// Mitsubishi GX Works2 project: 30国轩预化成10.29,排队位置优化   PLC: Q10UDEH

TYPE ConveyorIO : STRUCT
  xUnloadCCW : BOOL;  (* 下料为反转 *)
  xUnloadAlarm : BOOL;  (* 下料报警 *)
  xUnload : BOOL;  (* 下料请求 *)
  xPutInto : BOOL;  (* 线体直接投入物料 *)
  xNotArriveAlarm : BOOL;  (* 未到达报警 *)
  xNextRun : BOOL;  (* 下段线体运行 *)
  xMotorCW : BOOL;  (* 电机正转 *)
  xMotorCCW : BOOL;  (* 电机反转 *)
  xManual : BOOL;  (* 手动 *)
  xloadCCW : BOOL;  (* 上料为反转 *)
  xLimitAlarrm : BOOL;  (* 限位报警 *)
  xLoad : BOOL;  (* 上料请求 *)
  xForward : BOOL;  (* 正转手动 *)
  xEmpty : BOOL;  (* 线体状态为空 *)
  xCWPresent : BOOL;  (* 正转检测有无传感器 *)
  xCCWPresent : BOOL;  (* 反转检测有无传感器 *)
  xBusy : BOOL;  (* 工作中 *)
  xBackward : BOOL;  (* 反转手动 *)
  xAuto : BOOL;  (* 自动 *)
  xPosLimit : BOOL;  (* 正限位 *)
  xNegLimit : BOOL;  (* 负限位 *)
  xOverWidthAlarm : BOOL;  (* 超宽报警 *)
  xError : BOOL;  (* 报警 *)
  iProductCategoryIn : INT;  (* 产品类型输入 *)
  iProductCategory : INT;  (* 产品类型记录 *)
  iProductCategoryOut : INT;  (* 产品类型输出 *)
  diDeviceID : DINT;  (* 设备编号 *)
  tUnloadAlarmDelay : TIME;  (* 下料报警时间设置 *)
  tLoadDelay : TIME;  (* 上料延时设置 *)
  xSizeDeficientDetect : BOOL;  (* 尺寸缺陷检测 *)
  xZoneClear : BOOL;  (* 初始化线体清除 *)
  tZoneClearTime : TIME;  (* 初始化线体清除时间 *)
  iTaskIDIn : INT;  (* 产品类型输入 *)
  iTaskID : INT;  (* 产品类型记录 *)
  iTaskIDOut : INT;  (* 产品类型输出 *)
  diDesConveyorIn : DINT;  (* 产品类型输入 *)
  diDesConveyor : DINT;  (* 产品类型记录 *)
  diDesConveyorOut : DINT;  (* 产品类型输出 *)
END_STRUCT END_TYPE

TYPE ShuttleCarIO : STRUCT
  xReady : BOOL;  (* 准备就绪 *)
  xForward : BOOL;  (* 正转 *)
  xBackward : BOOL;  (* 反转 *)
  iCurrentPos : INT;  (* 当前位置 *)
  iDestinationPos : INT;  (* 目标位置 *)
  xCW : BOOL;  (* 正转输出 *)
  xCCW : BOOL;  (* 反转输出 *)
  xBrake : BOOL;  (* 刹车 *)
  xHomeSwitch : BOOL;  (* 零位接近开关 *)
  xPosLimit : BOOL;  (* 正限位 *)
  xNegLimit : BOOL;  (* 负限位 *)
  xMDIExe : BOOL;  (* MDI开始 *)
  xMDIDone : BOOL;  (* MDI 完成 *)
  xPassLimit : BOOL;  (* 限位屏蔽 *)
  xPosLimitCatch : BOOL;  (* 正限位捕捉 *)
  xNegLimitCatch : BOOL;  (* 负限位捕捉 *)
  xHomeExe : BOOL;  (* 开始寻零 *)
  xHomeDone : BOOL;  (* 寻零完成 *)
  xHomeBusy : BOOL;  (* 寻零中 *)
  xHomeFailed : BOOL;  (* 寻零失败 *)
  xBusy : BOOL;  (* 工作中 *)
  tArriveDelay : TIME;  (* 到位延时 *)
  xCylinder : BOOL;  (* 气缸控制 *)
  tBrakeDelay : TIME;  (* 抱闸延时 *)
  xPauseRamp : BOOL;  (* 暂停减速斜坡标志位 *)
  xPresentDetect1 : BOOL;  (* 物料有无检测1 *)
  xPresentDetect2 : BOOL;  (* 物料有无检测2 *)
  xOvertimeAlarm : BOOL;  (* 超时报警 *)
  tSetOverTime : TIME;  (* 设置超时时间 *)
  xLooseDetect : BOOL;  (* 松绳检测 *)
  xLooseAlarm : BOOL;  (* 松绳报警 *)
  xArrive : BOOL;  (* 到位信号 *)
  diDeviceID : DINT;  (* 设备编号 *)
  xMoveStep : BOOL;  (* 寸动 *)
  xAdrSwitch : ARRAY [1..8] OF BOOL;  (* 位置开关 *)
END_STRUCT END_TYPE

TYPE SwitchIO : STRUCT
  xLiftCylinderRetractDetect : BOOL;
  xLiftCylinderExtendDetect : BOOL;
  xLiftCylinderRetract : BOOL;
  xLiftCylinderExtend : BOOL;
  xEntryBarCylinderRetract : BOOL;
  xLiftCylinderExtendInit : BOOL;
  xEntryEnable : BOOL;
  xExitEnable : BOOL;
  xExitBarCylinderRetract : BOOL;
  xSwithEnable : BOOL;
  xLiftCylinderRetractButton : BOOL;
  xLiftCylinderExtendButton : BOOL;
  xEntryBarCylinderRetractButton : BOOL;
  xExitBarCylinderRetractButton : BOOL;
  xPutInto : BOOL;  (* 单体复位 *)
  tSetOvertime : TIME;  (* 设定超时报警时间 *)
  xOvertimeAlarm : BOOL;  (* 超时报警 *)
END_STRUCT END_TYPE

TYPE QueueElement : STRUCT
  xCondition : BOOL;
  iPriority : INT;
END_STRUCT END_TYPE

TYPE UConveyorIO : STRUCT
  xLiftCylinderRetractDetect1 : BOOL;
  xLiftCylinderRetractDetect2 : BOOL;
  xLiftCylinderExtendDetect1 : BOOL;
  xLiftCylinderExtendDetect2 : BOOL;
  xLiftCylinderRetract1 : BOOL;
  xLiftCylinderRetract2 : BOOL;
  xLiftCylinderExtend1 : BOOL;
  xLiftCylinderExtend2 : BOOL;
  xExitBarCylinderRetract1 : BOOL;
  xExitBarCylinderRetract2 : BOOL;
  xLiftCylinderExtendInit1 : BOOL;
  xLiftCylinderExtendInit2 : BOOL;
  xEntryEnable1 : BOOL;
  xEntryEnable2 : BOOL;
  xEntryEnable3 : BOOL;
  xExitEnable1 : BOOL;
  xExitEnable2 : BOOL;
  xExitEnable3 : BOOL;
  xPassEnable : BOOL;  (* 直接放行去下段 *)
  xLiftCylinderRetractButton1 : BOOL;
  xLiftCylinderRetractButton2 : BOOL;
  xLiftCylinderExtendButton1 : BOOL;
  xLiftCylinderExtendButton2 : BOOL;
  xExitBarCylinderRetractButton1 : BOOL;
  xExitBarCylinderRetractButton2 : BOOL;
  xPutInto : BOOL;  (* 单体复位 *)
  tSetOvertime : TIME;  (* 设定超时报警时间 *)
  xOvertimeAlarm : BOOL;  (* 超时报警 *)
  iTask : INT;  (* 3个任务 *)
  xBatteryDetect1 : BOOL;  (* 电池检测1 *)
  xBatteryDetect2 : BOOL;  (* 电池检测2 *)
  xBatteryError : BOOL;  (* 空框里有电池错误 *)
END_STRUCT END_TYPE

TYPE FolderIO : STRUCT
  o_xCylinderGrabExtend : BOOL;  (* 气缸夹紧 *)
  o_xCylinderGrabRetract : BOOL;  (* 气缸松开 *)
  i_xCylinderGrabExtendDetect : BOOL;  (* 夹紧检测 *)
  i_xCylinderGrabRetractDetect : BOOL;  (* 松开检测 *)
  o_xCylinderUpExtend : BOOL;  (* 上层伸出 *)
  o_xCylinderUpRetract : BOOL;  (* 上层缩回 *)
  i_xCylinderUpExtendDetect : BOOL;  (* 上层伸出检测 *)
  i_xCylinderUpRetractDetect : BOOL;  (* 上层缩回检测 *)
  o_xCylinderDownExtend : BOOL;  (* 下层伸出 *)
  o_xCylinderDownRetract : BOOL;  (* 下层缩回 *)
  i_xCylinderDownExtendDetect : BOOL;  (* 下层伸出检测 *)
  i_xCylinderDownRetractDetect : BOOL;  (* 下层缩回检测 *)
  i_xExitEnable : BOOL;  (* 下料信号 *)
  i_xEntryEnable : BOOL;  (* 上料信号 *)
  o_xEntryPermit : BOOL;  (* 允许上料 *)
  i_iFloor : INT;  (* 层数 *)
  i_xCylinderGrabExtendButton : BOOL;  (* 气缸夹紧按钮 *)
  i_xCylinderGrabRetractButton : BOOL;  (* 气缸松开按钮 *)
  i_xCylinderUpExtendButton : BOOL;  (* 上层伸出按钮 *)
  i_xCylinderUpRetractButton : BOOL;  (* 上层缩回按钮 *)
  i_xCylinderDownExtendButton : BOOL;  (* 下层伸出按钮 *)
  i_xCylinderDownRetractButton : BOOL;  (* 下层缩回按钮 *)
  o_xDownCylinderError : BOOL;  (* 下层气缸层伸出未到达 *)
  o_xUpCylinderError : BOOL;  (* 上层气缸伸出未到达 *)
  o_xGrabCylinderError : BOOL;  (* 夹紧气缸伸出未到达 *)
  i_tSetOvertime : TIME;  (* 未到达计时 *)
END_STRUCT END_TYPE

TYPE CommunicationIO : STRUCT
  i_iResponsPCPLC : INT;  (* 上位机写入-请求确认 *)
  i_iReadWriteFlagPCPLC : INT;  (* 上位机写入-读写标志位 *)
  i_iTaskProcessFlagPCPLC : INT;  (* 上位机写入-任务处理标志位 *)
  i_iCommandPCPLC : INT;  (* 上位机写入-命令字 *)
  i_iTaskIDPCPLC : INT;  (* 上位机写入-任务号 *)
  i_diDestinationDevicePCPLC : DINT;  (* 上位机写入-目标设备号 *)
  i_iProductIDPCPLC : INT;  (* 上位机写入-框码后4位 *)
  o_iRequestPLCPC : INT;  (* 上位机读取-请求状态 *)
  o_iReadWriteFlagPLCPC : INT;  (* 上位机读取-读写标志位 *)
  o_iDeviceStatusPLCPC : INT;  (* 上位机读取-设备状态 *)
  o_iTaskIDPLCPC : INT;  (* 上位机读取-任务号 *)
  o_iProductIDPLCPC : INT;  (* 上位机读取-框码后4位 *)
  i_iTypeInfoPCPLC : INT;  (* 上位机写入-批次标识，是否同批次 *)
  o_iForceInportPLCPC : INT;  (* 上位机读取-强制入库 *)
  o_iEmptyPLCPC : INT;  (* 上位机读取-有料状态 *)
  o_iFolderNumberPLCPC : INT;  (* 上位机读取-叠盘数量 *)
  i_xExtraCondition : BOOL;  (* 发送请求时的额外条件,比如需要升降到位 *)
  i_xExportConveyor : BOOL;  (* 线体是出库线体还是入库线体 *)
END_STRUCT END_TYPE

TYPE FanucRobotIO : STRUCT
  i_xCMDENBL : BOOL;
  i_xSYSRDY : BOOL;
  i_xPROG_RUN : BOOL;  (* 程序运行中 *)
  i_xPAUSED : BOOL;
  i_xHELD : BOOL;
  i_xFAULT : BOOL;
  i_xATPERCH : BOOL;
  i_xTPENBL : BOOL;
  i_xBATALM : BOOL;
  i_xBUSY : BOOL;  (* 工作中信号 *)
  i_arrxSNO : ARRAY [0..7] OF BOOL;  (* 传回的数据 *)
  i_xSNACK : BOOL;  (* 数据传回校验标志位 *)
  o_xIMSTP : BOOL;
  o_xHOLD : BOOL;
  o_xSFSPD : BOOL;
  o_xCSTOPI : BOOL;
  o_xRESET : BOOL;
  o_xSTART : BOOL;
  o_xENBL : BOOL;
  o_iPNS : INT;  (* 发给他的动作编号 *)
  o_xPNSTROBE : BOOL;  (* 传递动作编号标志位 *)
  o_xPROD_START : BOOL;  (* 启动信号，下降沿开动 *)
  o_xREMOTE : BOOL;  (* 远程模式开启 *)
  i_xCommandStart : BOOL;  (* 启动 *)
  i_iMotionNumber : INT;  (* 我程序给的动作编号 *)
  o_xPNSFailed : BOOL;  (* 程序号传输错误 *)
  o_uiOffset_X : INT;  (* X轴偏移量 *)
  o_uiOffset_Y : INT;  (* Y轴偏移量 *)
  io_xMutexLock : BOOL;  (* 互斥锁 *)
END_STRUCT END_TYPE

TYPE SortCommunicationIO : STRUCT
  i_iResponsPCPLC : INT;  (* 上位机写入-应答 *)
  i_iSortDoneAknPCPLC : INT;  (* 上位机写入-任务处理完成 *)
  i_arriBatteryStatus : ARRAY [1..128] OF INT;  (* 上位机写入-电池状态 *)
  o_iRequestPLCPC : INT;  (* 上位机读取-请求 *)
  o_iSortDonePLCPC : INT;  (* 上位机读取-分拣完成 *)
  i_iInfoWriteDone : INT;  (* 上位机写入-参数写入完成 *)
END_STRUCT END_TYPE

// global labels: Global
VAR_GLOBAL
  g_xAuto AT M11 : BOOL;
  g_xManual : BOOL;
  g_xEStop AT X0 : BOOL;
  g_xReset : BOOL;
  g_xStackLampRed AT Y200 : BOOL;  (* 塔灯红 *)
  g_xStackLampAmber AT Y201 : BOOL;  (* 塔灯黄 *)
  g_xStackLampGreen AT Y202 : BOOL;  (* 塔灯绿 *)
  g_xBuzzer AT Y203 : BOOL;  (* 蜂鸣器 *)
  g_xStop AT X3 : BOOL;
  g_xAutoStart AT X2 : BOOL;  (* 启动按钮 *)
  g_xRemoteAutoStart AT M0 : BOOL;
  g_xRemoteAuto AT M10 : BOOL;
  g_iState AT D40 : INT;  (* 状态显示 *)
  g_iLocalAutoStep : BOOL;
  g_xAlarm : BOOL;
  g_xPause AT M3 : BOOL;  (* 暂停 *)
  g_diDeviceIDSelect AT D0 : DINT;
  g_xResetSingle AT M4 : BOOL;  (* 单线体复位 *)
  g_xInsertTask AT M5 : BOOL;  (* 插入任务 *)
  g_iInsertTaskID AT D2 : INT;  (* 插入任务号 *)
  g_iConveyorStatus AT D4 : INT;
  g_iInsertCategory AT D6 : INT;
  g_diInsertDesConveyor AT D8 : DINT;
  g_x20TcpFailed : BOOL;  (* 30预20通讯失败 *)
  g_xAutoLamp AT Y204 : BOOL;  (* 启动灯 *)
  g_iLoadTask AT D50 : ARRAY [0..13] OF INT;  (* 排队任务站，D50-D62 *)
  g_xAutoSwitch AT X1 : BOOL;  (* 手自动钥匙旋钮 *)
  g_xMute AT M2 : BOOL;  (* 静音按钮，报警消除时复位 *)
  g_xResetTask1 AT M9 : BOOL;  (* 复位排队任务按钮 *)
  g_xLoadPermit : ARRAY [1..2] OF BOOL;  (* 定位机排队任务允许 *)
  g_x40TcpFailed : BOOL;  (* 30预40通讯失败 *)
  g_xForceImport AT M1 : BOOL;  (* 强制入库 *)
  g_x24HourImport1Forbidden AT M12 : BOOL;  (* 24小时入库禁止1 *)
  g_x24HourImport2Forbidden AT M13 : BOOL;  (* 24小时入库禁止2 *)
  g_xPreChemImport1Forbidden AT M14 : BOOL;  (* 预化成入库禁止1 *)
  g_xPreChemImport2Forbidden AT M15 : BOOL;  (* 预化成入库禁止2 *)
  g_x24HourExport1Forbidden AT M16 : BOOL;  (* 24小时出库禁止 *)
  g_xPreChemExport1Forbidden AT M17 : BOOL;  (* 预化成出库禁止1 *)
  g_xPreChemExport2Forbidden AT M18 : BOOL;  (* 预化成出库禁止2 *)
  g_xPickDone : BOOL;  (* 分拣完成 *)
  g_xPickOver AT X4 : BOOL;  (* 注液机给我们的信号，待定 *)
END_VAR

// task Task_01 (event TRUE, interval 0, priority 31): POU, START, TCP

PROGRAM POU
VAR
  Conveyor30101 : Conveyor;
  Conveyor30102 : Conveyor;
  Conveyor30103 : Conveyor;
  Conveyor30104 : Conveyor;
  Conveyor30105 : Conveyor;
  Conveyor30106 : Conveyor;
  Conveyor30107 : Conveyor;
  Conveyor30108 : Conveyor;
  Conveyor30109 : Conveyor;
  Conveyor30110 : Conveyor;
  Conveyor30111 : Conveyor;
  Conveyor30112 : Conveyor;
  Conveyor30113 : Conveyor;
  Conveyor30114 : Conveyor;
  Conveyor30115 : Conveyor;
  Conveyor30116 : Conveyor;
  Conveyor30117 : Conveyor;
  Conveyor30118 : Conveyor;
  Conveyor30119 : Conveyor;
  Conveyor30120 : Conveyor;
  Conveyor30121 : Conveyor;
  Conveyor30122 : Conveyor;
  Conveyor30123 : Conveyor;
  Conveyor30124 : Conveyor;
  Conveyor30125 : Conveyor;
  Conveyor30126 : Conveyor;
  Conveyor30127 : Conveyor;
  Conveyor30128 : Conveyor;
  Conveyor30129 : Conveyor;
  Conveyor30130 : Conveyor;
  Conveyor30131 : Conveyor;
  Conveyor30132 : Conveyor;
  Conveyor30133 : Conveyor;
  Conveyor30134 : Conveyor;
  Conveyor30135 : Conveyor;
  Conveyor30136 : Conveyor;
  Conveyor30137 : Conveyor;
  Conveyor301021 : Conveyor;  (* 高温入库升降门前停止位 *)
  Conveyor301071 : Conveyor;  (* 高温出库升降门前停止位 *)
  ConveyorIO30101 : ConveyorIO;
  ConveyorIO30102 : ConveyorIO;
  ConveyorIO30103 : ConveyorIO;
  ConveyorIO30104 : ConveyorIO;
  ConveyorIO30105 : ConveyorIO;
  ConveyorIO30106 : ConveyorIO;
  ConveyorIO30107 : ConveyorIO;
  ConveyorIO30108 : ConveyorIO;
  ConveyorIO30109 : ConveyorIO;
  ConveyorIO30110 : ConveyorIO;
  ConveyorIO30111 : ConveyorIO;
  ConveyorIO30112 : ConveyorIO;
  ConveyorIO30113 : ConveyorIO;
  ConveyorIO30114 : ConveyorIO;
  ConveyorIO30115 : ConveyorIO;
  ConveyorIO30116 : ConveyorIO;
  ConveyorIO30117 : ConveyorIO;
  ConveyorIO30118 : ConveyorIO;
  ConveyorIO30119 : ConveyorIO;
  ConveyorIO30120 : ConveyorIO;
  ConveyorIO30121 : ConveyorIO;
  ConveyorIO30122 : ConveyorIO;
  ConveyorIO30123 : ConveyorIO;
  ConveyorIO30124 : ConveyorIO;
  ConveyorIO30125 : ConveyorIO;
  ConveyorIO30126 : ConveyorIO;
  ConveyorIO30127 : ConveyorIO;
  ConveyorIO30128 : ConveyorIO;
  ConveyorIO30129 : ConveyorIO;
  ConveyorIO30130 : ConveyorIO;
  ConveyorIO30131 : ConveyorIO;
  ConveyorIO30132 : ConveyorIO;
  ConveyorIO30133 : ConveyorIO;
  ConveyorIO30134 : ConveyorIO;
  ConveyorIO30135 : ConveyorIO;
  ConveyorIO30136 : ConveyorIO;
  ConveyorIO30137 : ConveyorIO;
  ConveyorIO301021 : ConveyorIO;  (* 高温入库升降门前停止位 *)
  ConveyorIO301071 : ConveyorIO;  (* 高温出库升降门前停止位 *)
  Rotor30401 : ShuttleCar;
  Rotor30402 : ShuttleCar;
  Rotor30403 : ShuttleCar;
  Rotor30404 : ShuttleCar;
  Lifter30201 : ShuttleCar;
  Lifter30202 : ShuttleCar;
  Lifter30203 : ShuttleCar;
  Lifter30204 : ShuttleCar;
  Lifter30205 : ShuttleCar;
  Lifter30206 : ShuttleCar;
  Lifter30212 : ShuttleCar;
  Lifter30213 : ShuttleCar;
  Lifter30214 : ShuttleCar;
  Lifter30215 : ShuttleCar;
  RotorIO30401 : ShuttleCarIO;
  RotorIO30402 : ShuttleCarIO;
  RotorIO30403 : ShuttleCarIO;
  RotorIO30404 : ShuttleCarIO;
  LifterIO30201 : ShuttleCarIO;
  LifterIO30202 : ShuttleCarIO;
  LifterIO30203 : ShuttleCarIO;
  LifterIO30204 : ShuttleCarIO;
  LifterIO30205 : ShuttleCarIO;
  LifterIO30206 : ShuttleCarIO;
  LifterIO30212 : ShuttleCarIO;
  LifterIO30213 : ShuttleCarIO;
  LifterIO30214 : ShuttleCarIO;
  LifterIO30215 : ShuttleCarIO;
  Lifter30207 : ShuttleCar;
  LifterIO30207 : ShuttleCarIO;
  Switch30301 : Switch;
  Switch30302 : Switch;
  Switch30303 : Switch;
  Switch30304 : Switch;
  Switch30305 : Switch;
  Switch30306 : Switch;
  Switch30307 : Switch;
  Switch30308 : Switch;
  Switch30309 : Switch;
  Switch30310 : Switch;
  Switch30311 : Switch;
  SwitchIO30301 : SwitchIO;
  SwitchIO30302 : SwitchIO;
  SwitchIO30303 : SwitchIO;
  SwitchIO30304 : SwitchIO;
  SwitchIO30305 : SwitchIO;
  SwitchIO30306 : SwitchIO;
  SwitchIO30307 : SwitchIO;
  SwitchIO30308 : SwitchIO;
  SwitchIO30309 : SwitchIO;
  SwitchIO30310 : SwitchIO;
  SwitchIO30311 : SwitchIO;
  Conveyor301271 : Conveyor;
  ConveyorIO301271 : ConveyorIO;
  ConveyorIO30138 : ConveyorIO;
  ConveyorIO30139 : ConveyorIO;
  ConveyorIO30140 : ConveyorIO;
  Conveyor30138 : Conveyor;
  Conveyor30139 : Conveyor;
  Conveyor30140 : Conveyor;
  Conveyor301201 : Conveyor;
  ConveyorIO301201 : ConveyorIO;
  ComConveyor30103 : ConveyorCommunication;
  ComConveyor30136 : ConveyorCommunication;
  ComConveyor30104 : ConveyorCommunication;
  ComConveyor30137 : ConveyorCommunication;
  ComConveyor30111 : ConveyorCommunication;
  ComConveyor30116 : ConveyorCommunication;
  ComConveyor30112 : ConveyorCommunication;
  ComConveyor30117 : ConveyorCommunication;
  ComConveyor30114 : ConveyorCommunication;
  ComConveyor30119 : ConveyorCommunication;
  SortConveyor30121 : SortCommunication;
  ComConveyorIO30103 : CommunicationIO;
  ComConveyorIO30136 : CommunicationIO;
  ComConveyorIO30104 : CommunicationIO;
  ComConveyorIO30137 : CommunicationIO;
  ComConveyorIO30111 : CommunicationIO;
  ComConveyorIO30116 : CommunicationIO;
  ComConveyorIO30112 : CommunicationIO;
  ComConveyorIO30117 : CommunicationIO;
  ComConveyorIO30114 : CommunicationIO;
  ComConveyorIO30119 : CommunicationIO;
  SortConveyorIO30121 : SortCommunicationIO;
  Conveyor301111 : Conveyor;
  Conveyor301161 : Conveyor;
  ConveyorIO301111 : ConveyorIO;
  ConveyorIO301161 : ConveyorIO;
  Task30305 : PreemptivePriority;  (* 化成1巷道入库抢占任务 *)
  Task30305Condition : ARRAY [1..13] OF BOOL;  (* 化成1巷道入库抢占任务 *)
  m_iTask30305 : INT;  (* 化成1巷道入库抢占任务 *)
  Task30308 : PreemptivePriority;  (* 化成2巷道出库抢占任务 *)
  Task30308Condition : ARRAY [1..13] OF BOOL;  (* 化成2巷道出库抢占任务 *)
  m_iTask30308 : INT;  (* 化成2巷道出库抢占任务 *)
  Task30306 : PreemptivePriority;  (* 化成1巷道出库抢占任务 *)
  Task30306Condition : ARRAY [1..13] OF BOOL;  (* 化成1巷道出库抢占任务 *)
  m_iTask30306 : INT;  (* 化成1巷道出库抢占任务 *)
  Task30303 : PriorityQueue;  (* 化成12巷道入库任务分配 *)
  Task30303Condition : ARRAY [1..13] OF QueueElement;  (* 化成12巷道入库任务分配 *)
  m_iTask30303 : INT;  (* 化成12巷道入库任务分配 *)
  m_xRotor30401Start : BOOL;  (* 转台开始旋转 *)
  m_xRotor30402Start : BOOL;  (* 转台开始旋转 *)
  m_xRotor30403Start : BOOL;  (* 转台开始旋转 *)
  m_xRotor30404Start : BOOL;  (* 转台开始旋转 *)
  m_xRotor30401Done : BOOL;  (* 转台旋转完毕 *)
  m_xRotor30402Done : BOOL;  (* 转台旋转完毕 *)
  m_xRotor30403Done : BOOL;  (* 转台旋转完毕 *)
  m_xRotor30404Done : BOOL;  (* 转台旋转完毕 *)
  Conveyor30141 : Conveyor;
  Conveyor30142 : Conveyor;
  ConveyorIO30141 : ConveyorIO;
  ConveyorIO30142 : ConveyorIO;
  Conveyor301051 : Conveyor;  (* 高温出库后停止位 *)
  ConveyorIO301051 : ConveyorIO;  (* 高温出库后停止位 *)
  m_xLocation2Empty : BOOL;  (* 定位机2无料信号 *)
  m_xLocation1Load : BOOL;  (* 定位机1上料 *)
  m_xLocation2Load : BOOL;  (* 定位机2上料 *)
  m_xLocation1Unload : BOOL;  (* 定位机1下料 *)
  m_xLocation2Unload : BOOL;  (* 定位机2下料 *)
  m_xLocation1NextRun : BOOL;  (* 定位机1矫正完成 *)
  m_xLocation2NextRun : BOOL;  (* 定位机2矫正完成 *)
  m_xLocation1Empty : BOOL;  (* 定位机1无料信号 *)
  FanucRobotIO300 : FanucRobotIO;  (* 分拣机器人IO *)
  FanucRobot300 : FanucRobot;  (* 分拣机器人 *)
END_VAR
(*和定位机对接信号*)
Y23D:=m_xLocation1Load;(*定位机上料中，我们发给他的，让他转起来上料*)
Y23F:=m_xLocation1Unload;(*定位机下料中，我们发给他的，让他转起来下料*)
m_xLocation1Empty:=X7D;(*定位机为空，给我们上料请求*)
m_xLocation1NextRun:=X7F;(*定位机定位完，给我们的下料请求*)

Y241:=m_xLocation2Load;(*定位机上料中，我们发给他的，让他转起来上料*)
Y243:=m_xLocation2Unload;(*定位机下料中，我们发给他的，让他转起来下料*)
m_xLocation2Empty:=X81;(*定位机为空，给我们上料请求*)
m_xLocation2NextRun:=X83;(*定位机定位完，给我们的下料请求*)

Conveyor30101(ConveyorMotor:=ConveyorIO30101);(*高温库入库横向*)
ConveyorIO30101.xCWPresent:=X8;						
Y208:=ConveyorIO30101.xMotorCW;						
ConveyorIO30101.xForward:=M500;						
M301:= NOT ConveyorIO30101.xEmpty;						
M601:=ConveyorIO30101.xError;						
ConveyorIO30101.diDeviceID:=30101;	
ConveyorIO30101.tLoadDelay:=t#400ms;

Conveyor30102(ConveyorMotor:=ConveyorIO30102);
ConveyorIO30102.xCCWPresent:=X8;(*01和02组成switch，高温入库门前的*)
Y209:=ConveyorIO30102.xMotorCW OR ConveyorIO301021.xMotorCW ;						
ConveyorIO30102.xForward:=M501;														
M602:=ConveyorIO30102.xError OR ConveyorIO301021.xError;						
ConveyorIO30102.diDeviceID:=301021;			
			
Conveyor301021(ConveyorMotor:=ConveyorIO301021);
ConveyorIO301021.xCWPresent:=X9;(*门前停止位，要虚拟一段线体*)								
M302:= NOT ConveyorIO301021.xEmpty;											
ConveyorIO301021.diDeviceID:=30102;			
			
Conveyor30103(ConveyorMotor:=ConveyorIO30103);(*高温库入库门后竖向线体*)
ConveyorIO30103.xCWPresent:=XA;						
Y20A:=ConveyorIO30103.xMotorCW;						
ConveyorIO30103.xForward:=M502;						
M303:= NOT ConveyorIO30103.xEmpty;
M603:=ConveyorIO30103.xError;
ConveyorIO30103.diDeviceID:=30103;		
ConveyorIO30103.tLoadDelay:=t#4500MS;

Conveyor30141(ConveyorMotor:=ConveyorIO30141);
ConveyorIO30141.xCWPresent:=XA;		(*41和03组成switch，入库门后那个*)				
Y21E:=ConveyorIO30141.xMotorCW;						
ConveyorIO30141.xForward:=M586;	
M341:=NOT ConveyorIO30141.xEmpty;
M641:=ConveyorIO30141.xError;						
ConveyorIO30141.diDeviceID:=30141;	

Conveyor30104(ConveyorMotor:=ConveyorIO30104);(*高温库入库对接*)
ConveyorIO30104.xCWPresent:=XB;						
Y20B:=ConveyorIO30104.xMotorCW;						
ConveyorIO30104.xForward:=M503;						
M304:= NOT ConveyorIO30104.xEmpty;						
M604:=ConveyorIO30104.xError;						
ConveyorIO30104.diDeviceID:=30104;						
ConveyorIO30104.tLoadDelay:=t#6500ms;

Conveyor30136(ConveyorMotor:=ConveyorIO30136);
(*ConveyorIO30136.xPosLimit:=XA2*);	(*04后的一段，入库对接，开始以为是一段，就没写*)					
ConveyorIO30136.xCWPresent:=XA6;			
Y27A:=ConveyorIO30136.xMotorCW;
ConveyorIO30136.xForward:=M587;
M336:= NOT ConveyorIO30136.xEmpty;						
M636:=ConveyorIO30136.xError;						
ConveyorIO30136.diDeviceID:=30136;
ConveyorIO30136.tLoadDelay:=t#1000ms;	

Conveyor30109(ConveyorMotor:=ConveyorIO30109);(*高温库出库对接*)
ConveyorIO30109.xCWPresent:=X10;						
Y210:=ConveyorIO30109.xMotorCW;						
ConveyorIO30109.xForward:=M508;						
M309:= NOT ConveyorIO30109.xEmpty;						
M609:=ConveyorIO30109.xError;						
ConveyorIO30109.diDeviceID:=30109;						
ConveyorIO30109.tLoadDelay:=t#6500ms;
Conveyor30137(ConveyorMotor:=ConveyorIO30137);	(*09前面末端那个线体，高温库出库对接*)				
ConveyorIO30137.xCWPresent:=XA3;
Y27B:=ConveyorIO30137.xMotorCW;
ConveyorIO30137.xForward:=M589;
M337:= NOT ConveyorIO30137.xEmpty;						
M637:=ConveyorIO30137.xError;						
ConveyorIO30137.diDeviceID:=30137;					

Conveyor30142(ConveyorMotor:=ConveyorIO30142);
ConveyorIO30142.xCWPresent:=XA7;			(*和08组成switch，横向*)			
Y21C:=ConveyorIO30142.xMotorCW;						
ConveyorIO30142.xForward:=M588;						
M342:= NOT ConveyorIO30142.xEmpty;						
M642:=ConveyorIO30142.xError;						
ConveyorIO30142.diDeviceID:=30142;	
ConveyorIO30142.tLoadDelay:=t#5000ms;	

Conveyor30108(ConveyorMotor:=ConveyorIO30108);(*高温出库门后switch，竖向线体*)
ConveyorIO30108.xCWPresent:=XA7;											
Y20F:=ConveyorIO30108.xMotorCW OR ConveyorIO301071.xMotorCW;						
ConveyorIO30108.xForward:=M507;					
M608:=ConveyorIO30108.xError OR ConveyorIO301071.xError;						
ConveyorIO30108.diDeviceID:=301071;		

Conveyor301071(ConveyorMotor:=ConveyorIO301071);
ConveyorIO301071.xCWPresent:=XF;		(*08到门前停止位，虚拟的*)										
M308:= NOT ConveyorIO301071.xEmpty;	
ConveyorIO301071.diDeviceID:=30108;

Conveyor30107(ConveyorMotor:=ConveyorIO30107);
ConveyorIO30107.xCWPresent:=XC;		(*07和05组成一个switch*)				
Y20E:=ConveyorIO30107.xMotorCW;						
ConveyorIO30107.xForward:=M506;						
M307:= NOT ConveyorIO30107.xEmpty;						
M607:=ConveyorIO30107.xError;						
ConveyorIO30107.diDeviceID:=30107;	
ConveyorIO30107.tLoadDelay:=t#3000ms;

Conveyor30105(ConveyorMotor:=ConveyorIO30105);(*高温出库横向线体，和07组成switch*)
ConveyorIO30105.xCWPresent:=XC;	
Y20C:=ConveyorIO30105.xMotorCW OR ConveyorIO301051.xMotorCW;						
ConveyorIO30105.xForward:=M504;																
M605:=ConveyorIO30105.xError OR ConveyorIO301051.xError;						
ConveyorIO30105.diDeviceID:=30105;						

Conveyor301051(ConveyorMotor:=ConveyorIO301051);(*高温出库后05后面，需要停在化成入库前，所以虚拟一段*)
ConveyorIO301051.xCWPresent:=XD;												
M305:= NOT ConveyorIO301051.xEmpty;							
ConveyorIO301051.diDeviceID:=30105;										

Conveyor30106(ConveyorMotor:=ConveyorIO30106);(*预化成1入库横向线体，和11组成switch*)
ConveyorIO30106.xCWPresent:=X2F;						
Y20D:=ConveyorIO30106.xMotorCW;						
ConveyorIO30106.xForward:=M505;						
M306:= NOT ConveyorIO30106.xEmpty;						
M606:=ConveyorIO30106.xError;						
ConveyorIO30106.diDeviceID:=30106;
ConveyorIO30106.tLoadDelay:=t#7500ms;

Conveyor30111(ConveyorMotor:=ConveyorIO30111);(*和06组成switch*)
ConveyorIO30111.xCWPresent:=X2F;	
Y212:=ConveyorIO301111.xMotorCW OR ConveyorIO30111.xMotorCW;	
ConveyorIO301111.xForward:=M510;													
M311:= NOT ConveyorIO30111.xEmpty;						
M611:=ConveyorIO30111.xError;						
ConveyorIO30111.diDeviceID:=30111;						
ConveyorIO30111.tLoadDelay:=t#4000ms;

Conveyor301111(ConveyorMotor:=ConveyorIO301111);(*化成1入库门前停止位，虚拟一段,暂时取消由定位机代替了*)
ConveyorIO301111.xCWPresent:=X12;		

Conveyor30134(ConveyorMotor:=ConveyorIO30134);(*预化成1入库转台线体*)
ConveyorIO30134.xPosLimit:=NOT X71;						
ConveyorIO30134.xCWPresent:=X70;						
Y269:=ConveyorIO30134.xMotorCW;			
Y268:=ConveyorIO30134.xMotorCCW;			
ConveyorIO30134.xForward:=M535;	
ConveyorIO30134.xBackward:=M590;					
M334:= NOT ConveyorIO30134.xEmpty;						
M634:=ConveyorIO30134.xError;						
ConveyorIO30134.diDeviceID:=30134;						
Y24A:=ConveyorIO30134.xNextRun OR (g_xManual AND M595);	(*转台阻挡*)
ConveyorIO30134.tLoadDelay:=t#1S;

Conveyor30112(ConveyorMotor:=ConveyorIO30112);(*预化成入库对接线体*)
ConveyorIO30112.xCWPresent:=X13;			
ConveyorIO30112.xNegLimit:=XBD;
Y213:=ConveyorIO30112.xMotorCW;						
ConveyorIO30112.xForward:=M511;						
M312:= NOT ConveyorIO30112.xEmpty;						
M612:=ConveyorIO30112.xError;						
ConveyorIO30112.diDeviceID:=30112;	
ConveyorIO30112.tLoadDelay:=t#300ms;

Conveyor30114(ConveyorMotor:=ConveyorIO30114);(*预化成1出库对接线体*)
ConveyorIO30114.xCWPresent:=X15;
ConveyorIO30114.xCCWPresent:=XB1;
Y215:=ConveyorIO30114.xMotorCW;						
ConveyorIO30114.xForward:=M513;						
M314:= NOT ConveyorIO30114.xEmpty;						
M614:=ConveyorIO30114.xError;						
ConveyorIO30114.diDeviceID:=30114;		

Conveyor30113(ConveyorMotor:=ConveyorIO30113);(*预化成1出库，和10组成switch*)
ConveyorIO30113.xCWPresent:=X11;					
Y214:=ConveyorIO30113.xMotorCW;						
ConveyorIO30113.xForward:=M512;						
M313:= NOT ConveyorIO30113.xEmpty;						
M613:=ConveyorIO30113.xError;						
ConveyorIO30113.diDeviceID:=30113;	
ConveyorIO30113.tLoadDelay:=t#4000ms;

Conveyor30110(ConveyorMotor:=ConveyorIO30110);(*预化成1出库横向线体，和13组成switch*)
ConveyorIO30110.xCWPresent:=X11;						
Y275:=ConveyorIO30110.xMotorCW OR ConveyorIO30138.xMotorCW ;						
ConveyorIO30110.xForward:=M509;										
ConveyorIO30110.diDeviceID:=30110;		
ConveyorIO30110.tLoadDelay:=t#4000ms;

Conveyor30138(ConveyorMotor:=ConveyorIO30138);(*10下一段，12库之间的过渡线体*)
ConveyorIO30138.xCWPresent:=XB5;											
M310:= NOT ConveyorIO30138.xEmpty;						
M610:=ConveyorIO30138.xError;						
ConveyorIO30138.diDeviceID:=30110;															

Conveyor30115(ConveyorMotor:=ConveyorIO30115);(*预化成2入库横向线体*)
ConveyorIO30115.xCWPresent:=X16;						
Y216:=ConveyorIO30115.xMotorCW;						
ConveyorIO30115.xForward:=M514;						
M315:= NOT ConveyorIO30115.xEmpty;						
M615:=ConveyorIO30115.xError;						
ConveyorIO30115.diDeviceID:=30115;						
ConveyorIO30115.tLoadDelay:=t#4500ms;

Conveyor30116(ConveyorMotor:=ConveyorIO30116);(*预化成2入库竖向，和15组成switch*)
ConveyorIO30116.xCWPresent:=X16;	
Y217:=ConveyorIO30116.xMotorCW OR ConveyorIO301161.xMotorCW;						
ConveyorIO30116.xForward:=M515;									
M316:= NOT ConveyorIO30116.xEmpty;						
M616:=ConveyorIO30116.xError;						
ConveyorIO30116.diDeviceID:=30116;						

Conveyor301161(ConveyorMotor:=ConveyorIO301161);(*门前停止位，虚拟线体，取消，由定位机代替*)
ConveyorIO301161.xCWPresent:=X17;	
ConveyorIO301161.diDeviceID:=301161;

Conveyor30117(ConveyorMotor:=ConveyorIO30117);(*预化成2入库对接线体*)
ConveyorIO30117.xNegLimit:=NOT XB2;
ConveyorIO30117.xCWPresent:=X18;						
Y218:=ConveyorIO30117.xMotorCW;						
ConveyorIO30117.xForward:=M516;						
M317:= NOT ConveyorIO30117.xEmpty;						
M617:=ConveyorIO30117.xError;						
ConveyorIO30117.diDeviceID:=30117;						

Conveyor30119(ConveyorMotor:=ConveyorIO30119);(*预化成2出库对接线体*)
ConveyorIO30119.xCWPresent:=X1A OR XB3;						
Y21A:=ConveyorIO30119.xMotorCW;						
ConveyorIO30119.xForward:=M518;						
M319:= NOT ConveyorIO30119.xEmpty;						
M619:=ConveyorIO30119.xError;						
ConveyorIO30119.diDeviceID:=30119;			

Conveyor30118(ConveyorMotor:=ConveyorIO30118);(*预化成2出库，和22组成switch*)
ConveyorIO30118.xCWPresent:=X9E;				
Y219:=ConveyorIO30118.xMotorCW;						
ConveyorIO30118.xForward:=M517;						
M318:= NOT ConveyorIO30118.xEmpty;						
M618:=ConveyorIO30118.xError;						
ConveyorIO30118.diDeviceID:=30118;		
ConveyorIO30118.tLoadDelay:=t#4000ms;							

Conveyor30122(ConveyorMotor:=ConveyorIO30122);(*预化成2出库横向线体，和18组成switch*)
ConveyorIO30122.xCWPresent:=X9E;						
Y21B:=ConveyorIO30122.xMotorCW;			
ConveyorIO30122.xForward:=M520;						
M322:= NOT ConveyorIO30122.xEmpty;						
M622:=ConveyorIO30122.xError;						
ConveyorIO30122.diDeviceID:=30122;	
(*图里是机械手用的线体，实际没有
Conveyor30120(ConveyorMotor:=ConveyorIO30120);
ConveyorIO30120.xCWPresent:=X1C;	
M320:= NOT ConveyorIO30120.xEmpty;						
M620:=ConveyorIO30120.xError;						
ConveyorIO30120.diDeviceID:=30120;						
*)
Conveyor30121(ConveyorMotor:=ConveyorIO30121);(*挑选机械手那段线体*)
ConveyorIO30121.xCWPresent:=X1E;						
Y21D:=ConveyorIO30121.xMotorCW;						
ConveyorIO30121.xForward:=M519;						
M321:= NOT ConveyorIO30121.xEmpty;						
M621:=ConveyorIO30121.xError;						
ConveyorIO30121.diDeviceID:=30121;										

Conveyor30123(ConveyorMotor:=ConveyorIO30123);
ConveyorIO30123.xCWPresent:=X20;						
Y21F:=ConveyorIO30123.xMotorCW;						
ConveyorIO30123.xForward:=M521;						
M323:= NOT ConveyorIO30123.xEmpty;						
M623:=ConveyorIO30123.xError;						
ConveyorIO30123.diDeviceID:=30123;						

Conveyor30124(ConveyorMotor:=ConveyorIO30124);(*下层1*)
ConveyorIO30124.xCWPresent:=X21;						
Y220:=ConveyorIO30124.xMotorCW;						
ConveyorIO30124.xForward:=M522;						
M324:= NOT ConveyorIO30124.xEmpty;						
M624:=ConveyorIO30124.xError;						
ConveyorIO30124.diDeviceID:=30124;						

Conveyor30125(ConveyorMotor:=ConveyorIO30125);(*下层2*)
ConveyorIO30125.xCWPresent:=X22;						
Y221:=ConveyorIO30125.xMotorCW;						
ConveyorIO30125.xForward:=M523;						
M325:= NOT ConveyorIO30125.xEmpty;						
M625:=ConveyorIO30125.xError;						
ConveyorIO30125.diDeviceID:=30125;						

Conveyor30126(ConveyorMotor:=ConveyorIO30126);(*下层3*)
ConveyorIO30126.xCWPresent:=X26;						
Y225:=ConveyorIO30126.xMotorCW;						
ConveyorIO30126.xForward:=M524;						
M326:= NOT ConveyorIO30126.xEmpty;						
M626:=ConveyorIO30126.xError;						
ConveyorIO30126.diDeviceID:=30126;						

Conveyor30127(ConveyorMotor:=ConveyorIO30127);
ConveyorIO30127.xCWPresent:=X26;						
Y226:=ConveyorIO30127.xMotorCW;						
Y223:=ConveyorIO30127.xMotorCCW;						
ConveyorIO30127.xForward:=M525;						
ConveyorIO30127.xBackward:=M526;						
M327:= NOT ConveyorIO30127.xEmpty;						
M627:=ConveyorIO30127.xError;						
ConveyorIO30127.diDeviceID:=30127;						

Conveyor30128(ConveyorMotor:=ConveyorIO30128);
ConveyorIO30128.xCWPresent:=X28;						
Y227:=ConveyorIO30128.xMotorCW;						
Y224:=ConveyorIO30128.xMotorCCW;						
ConveyorIO30128.xForward:=M527;						
ConveyorIO30128.xBackward:=M528;						
M328:= NOT ConveyorIO30128.xEmpty;						
M628:=ConveyorIO30128.xError;						
ConveyorIO30128.diDeviceID:=30128;						

Conveyor30129(ConveyorMotor:=ConveyorIO30129);
ConveyorIO30129.xCWPresent:=X25;						
ConveyorIO30129.xCCWPresent:=X29;						
Y274:=ConveyorIO30129.xMotorCW;						
Y276:=ConveyorIO30129.xMotorCCW;						
ConveyorIO30129.xForward:=M529;						
ConveyorIO30129.xBackward:=M530;						
M329:= NOT ConveyorIO30129.xEmpty;						
M629:=ConveyorIO30129.xError;						
ConveyorIO30129.diDeviceID:=30129;						

Conveyor30130(ConveyorMotor:=ConveyorIO30130);(*下层4*)
ConveyorIO30130.xCWPresent:=X23;
OUT_T( ConveyorIO30130.xMotorCW , TC0, 10);						
Y211:=TS0;						
ConveyorIO30130.xForward:=M531;						
M330:= NOT ConveyorIO30130.xEmpty;						
M630:=ConveyorIO30130.xError;						
ConveyorIO30130.diDeviceID:=30130;						

Conveyor30131(ConveyorMotor:=ConveyorIO30131);
ConveyorIO30131.xNegLimit:=NOT X77;						
ConveyorIO30131.xCWPresent:=X76;						
Y26F:=ConveyorIO30131.xMotorCW;
Y26E:=ConveyorIO30131.xMotorCCW;
ConveyorIO30131.xForward:=M532;
ConveyorIO30131.xBackward:=M593;							
M331:= NOT ConveyorIO30131.xEmpty;						
M631:=ConveyorIO30131.xError;						
ConveyorIO30131.diDeviceID:=30131;	
Y24C:=ConveyorIO30131.xNextRun OR  M598;	(*转台阻挡*)					

Conveyor30132(ConveyorMotor:=ConveyorIO30132);
ConveyorIO30132.xPosLimit:=NOT X75;						
ConveyorIO30132.xCWPresent:=X74;						
Y26C:=ConveyorIO30132.xMotorCW;
Y26D:=ConveyorIO30132.xMotorCCW;						
ConveyorIO30132.xForward:=M533;	
ConveyorIO30132.xBackward:=M592;						
M332:= NOT ConveyorIO30132.xEmpty;						
M632:=ConveyorIO30132.xError;						
ConveyorIO30132.diDeviceID:=30132;	
ConveyorIO30132.tLoadDelay:=t#1s;
Y24B:=ConveyorIO30132.xNextRun OR M597;	(*转台阻挡*)					

Conveyor30133(ConveyorMotor:=ConveyorIO30133);(*预化成1出库转台线体*)
ConveyorIO30133.xPosLimit:=(NOT X14 AND  NOT ConveyorIO30133.xUnloadCCW)OR ConveyorIO30133.xUnloadCCW ;	(*正转下料，这个开关作为正限位*)		
ConveyorIO30133.xNegLimit:=(NOT X14 AND ConveyorIO30133.xUnloadCCW)OR NOT ConveyorIO30133.xUnloadCCW ;	(*正转下料，这个开关作为正限位*)	
ConveyorIO30133.xCWPresent:=X72;						
Y26B:=ConveyorIO30133.xMotorCW;	
Y26A:=ConveyorIO30133.xMotorCCW;					
ConveyorIO30133.xForward:=M534;
ConveyorIO30133.xBackward:=M591;						
M333:= NOT ConveyorIO30133.xEmpty;						
M633:=ConveyorIO30133.xError;						
ConveyorIO30133.diDeviceID:=30133;	
ConveyorIO30133.tLoadDelay:=t#100MS;
Y249:=ConveyorIO30133.xNextRun OR (g_xManual AND M596);	(*转台阻挡*)

Conveyor30135(ConveyorMotor:=ConveyorIO30135);
ConveyorIO30135.xPosLimit:=NOT XA5;						
ConveyorIO30135.xCWPresent:=XA1;						
ConveyorIO30135.xCCWPresent:=XA4;						
Y278:=ConveyorIO30135.xMotorCW;						
Y279:=ConveyorIO30135.xMotorCCW;						
ConveyorIO30135.xForward:=M536;						
ConveyorIO30135.xBackward:=M537;						
M335:= NOT ConveyorIO30135.xEmpty;						
M635:=ConveyorIO30135.xError;						
ConveyorIO30135.diDeviceID:=30135;																				

Conveyor301271(ConveyorMotor:=ConveyorIO301271);
ConveyorIO301271.xCWPresent:=X28;						
M340:= NOT ConveyorIO301271.xEmpty;						
M640:=ConveyorIO301271.xError;						
ConveyorIO301271.diDeviceID:=301271;						

Conveyor30139(ConveyorMotor:=ConveyorIO30139);
ConveyorIO30139.xCWPresent:=X1C;						
Y27D:=ConveyorIO30139.xMotorCW;						
ConveyorIO30139.xForward:=M539;						
M339:= NOT ConveyorIO30139.xEmpty;						
M639:=ConveyorIO30139.xError;						
ConveyorIO30139.diDeviceID:=30139;						

Conveyor30140(ConveyorMotor:=ConveyorIO30140);
ConveyorIO30140.xCWPresent:=XB7 AND 0;		(**回流入库先屏蔽掉*)				
Y27E:=ConveyorIO30140.xMotorCW;						
ConveyorIO30140.xForward:=M540;						
M343:= NOT ConveyorIO30140.xEmpty;						
M643:=ConveyorIO30140.xError;						
ConveyorIO30140.diDeviceID:=30140;						